// TIA Portal project "FORMING_1500_PLC" (V15) (continued)
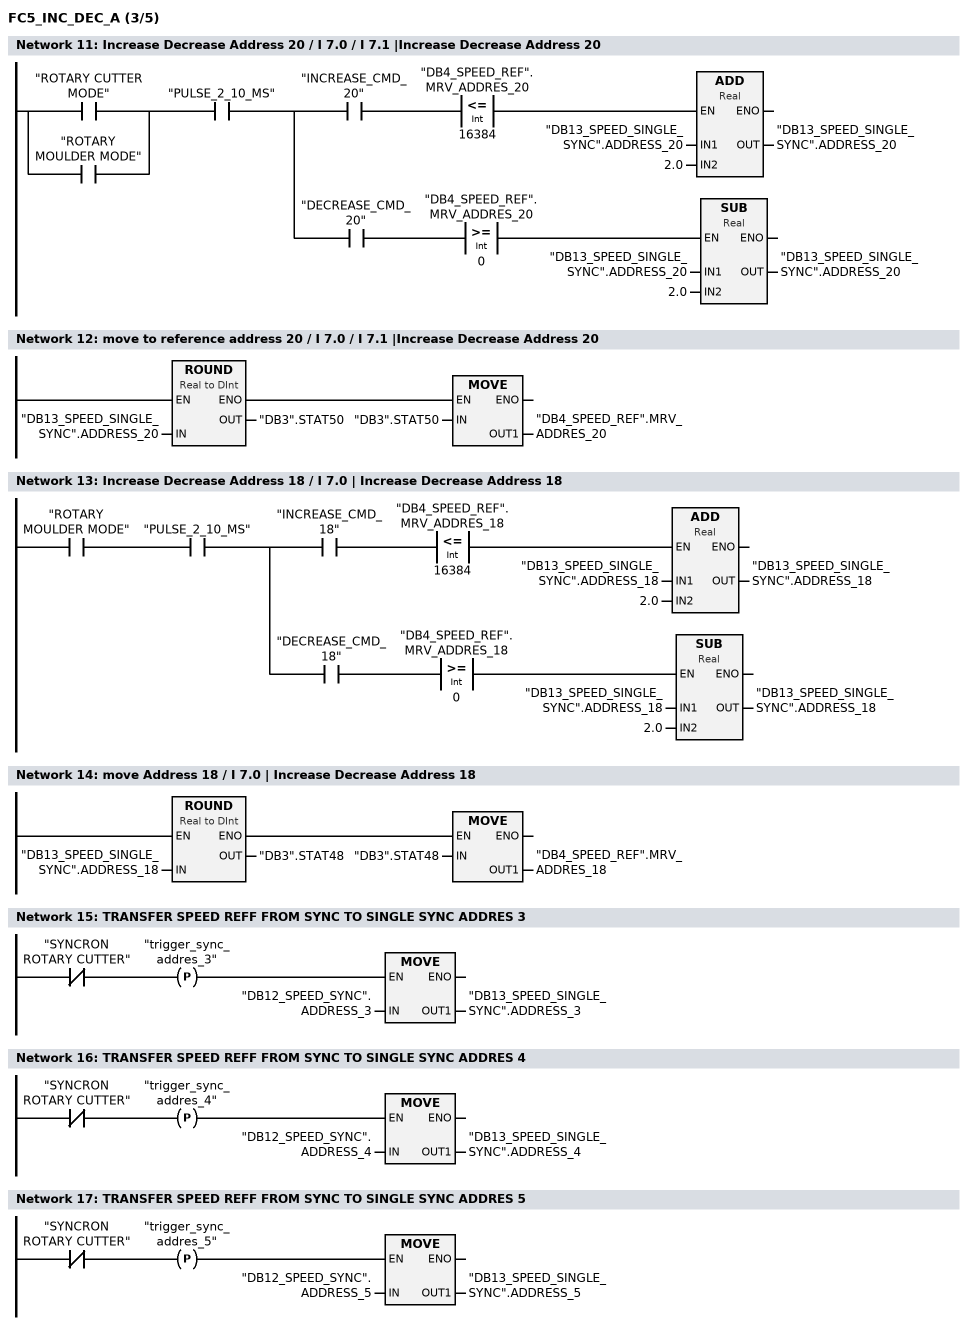
   RUNG wire#powerrail
      Contact( "ROTARY CUTTER MODE" )
      wire#w1
      Contact( "PULSE_2_10_MS" )
      wire#w2
      Contact( "INCREASE_CMD_20" )
      { S7_Templates := "SrcType := Int" } LE_Contact(in1 := "DB4_SPEED_REF".MRV_ADDRES_20, in2 := 16384)
      { S7_Templates := "SrcType := Real"; S7_GenerateENO := "TRUE" } Add(in1 := "DB13_SPEED_SINGLE_SYNC".ADDRESS_20, in2 := 2.0, out => "DB13_SPEED_SINGLE_SYNC".ADDRESS_20)
   END_RUNG
   RUNG wire#powerrail
      Contact( "ROTARY MOULDER MODE" )
   END_RUNG wire#w1
   RUNG wire#w2
      Contact( "DECREASE_CMD_20" )
      { S7_Templates := "SrcType := Int" } GE_Contact(in1 := "DB4_SPEED_REF".MRV_ADDRES_20, in2 := 0)
      { S7_Templates := "SrcType := Real"; S7_GenerateENO := "TRUE" } Sub(in1 := "DB13_SPEED_SINGLE_SYNC".ADDRESS_20, in2 := 2.0, out => "DB13_SPEED_SINGLE_SYNC".ADDRESS_20)
   END_RUNG
   // the same network as SCL:
   #_w1 := ("ROTARY CUTTER MODE" OR "ROTARY MOULDER MODE") AND "PULSE_2_10_MS";
   IF #_w1 AND "INCREASE_CMD_20" AND ("DB4_SPEED_REF".MRV_ADDRES_20 <= 16384) THEN
       "DB13_SPEED_SINGLE_SYNC".ADDRESS_20 := "DB13_SPEED_SINGLE_SYNC".ADDRESS_20 + 2.0;
   END_IF;
   IF #_w1 AND "DECREASE_CMD_20" AND ("DB4_SPEED_REF".MRV_ADDRES_20 >= 0) THEN
       "DB13_SPEED_SINGLE_SYNC".ADDRESS_20 := "DB13_SPEED_SINGLE_SYNC".ADDRESS_20 - 2.0;
   END_IF;
END_REGION

REGION Network 12: move to reference address 20 / I 7.0 / I 7.1 |Increase Decrease Address 20
   RUNG wire#powerrail
      { S7_Templates := "[SrcType := Real, DestType := DInt]"; S7_GenerateENO := "TRUE" } Round(in := "DB13_SPEED_SINGLE_SYNC".ADDRESS_20, out => "DB3".STAT50)
      { S7_GenerateENO := "TRUE" } Move(in := "DB3".STAT50, out1 => "DB4_SPEED_REF".MRV_ADDRES_20)
   END_RUNG
   // the same network as SCL:
   // ENO of a box is taken as its EN; it also drops when the box reports an error
   "DB3".STAT50 := ROUND("DB13_SPEED_SINGLE_SYNC".ADDRESS_20);
   "DB4_SPEED_REF".MRV_ADDRES_20 := "DB3".STAT50;
END_REGION

REGION Network 13: Increase Decrease Address 18 / I 7.0 | Increase Decrease Address 18
   RUNG wire#powerrail
      Contact( "ROTARY MOULDER MODE" )
      Contact( "PULSE_2_10_MS" )
      wire#w1
      Contact( "INCREASE_CMD_18" )
      { S7_Templates := "SrcType := Int" } LE_Contact(in1 := "DB4_SPEED_REF".MRV_ADDRES_18, in2 := 16384)
      { S7_Templates := "SrcType := Real"; S7_GenerateENO := "TRUE" } Add(in1 := "DB13_SPEED_SINGLE_SYNC".ADDRESS_18, in2 := 2.0, out => "DB13_SPEED_SINGLE_SYNC".ADDRESS_18)
   END_RUNG
   RUNG wire#w1
      Contact( "DECREASE_CMD_18" )
      { S7_Templates := "SrcType := Int" } GE_Contact(in1 := "DB4_SPEED_REF".MRV_ADDRES_18, in2 := 0)
      { S7_Templates := "SrcType := Real"; S7_GenerateENO := "TRUE" } Sub(in1 := "DB13_SPEED_SINGLE_SYNC".ADDRESS_18, in2 := 2.0, out => "DB13_SPEED_SINGLE_SYNC".ADDRESS_18)
   END_RUNG
   // the same network as SCL:
   #_w1 := "ROTARY MOULDER MODE" AND "PULSE_2_10_MS";
   IF #_w1 AND "INCREASE_CMD_18" AND ("DB4_SPEED_REF".MRV_ADDRES_18 <= 16384) THEN
       "DB13_SPEED_SINGLE_SYNC".ADDRESS_18 := "DB13_SPEED_SINGLE_SYNC".ADDRESS_18 + 2.0;
   END_IF;
   IF #_w1 AND "DECREASE_CMD_18" AND ("DB4_SPEED_REF".MRV_ADDRES_18 >= 0) THEN
       "DB13_SPEED_SINGLE_SYNC".ADDRESS_18 := "DB13_SPEED_SINGLE_SYNC".ADDRESS_18 - 2.0;
   END_IF;
END_REGION

REGION Network 14: move Address 18 / I 7.0 | Increase Decrease Address 18
   RUNG wire#powerrail
      { S7_Templates := "[SrcType := Real, DestType := DInt]"; S7_GenerateENO := "TRUE" } Round(in := "DB13_SPEED_SINGLE_SYNC".ADDRESS_18, out => "DB3".STAT48)
      { S7_GenerateENO := "TRUE" } Move(in := "DB3".STAT48, out1 => "DB4_SPEED_REF".MRV_ADDRES_18)
   END_RUNG
   // the same network as SCL:
   // ENO of a box is taken as its EN; it also drops when the box reports an error
   "DB3".STAT48 := ROUND("DB13_SPEED_SINGLE_SYNC".ADDRESS_18);
   "DB4_SPEED_REF".MRV_ADDRES_18 := "DB3".STAT48;
END_REGION

REGION Network 15: TRANSFER SPEED REFF FROM SYNC TO SINGLE SYNC ADDRES 3
   RUNG wire#powerrail
      I_Contact( "SYNCRON ROTARY CUTTER" )
      P_Trig( "trigger_sync_addres_3" )
      { S7_GenerateENO := "TRUE" } Move(in := "DB12_SPEED_SYNC".ADDRESS_3, out1 => "DB13_SPEED_SINGLE_SYNC".ADDRESS_3)
   END_RUNG
   // the same network as SCL:
   #_w1 := NOT "SYNCRON ROTARY CUTTER" AND NOT "trigger_sync_addres_3";   // rising edge
   "trigger_sync_addres_3" := NOT "SYNCRON ROTARY CUTTER";
   IF #_w1 THEN "DB13_SPEED_SINGLE_SYNC".ADDRESS_3 := "DB12_SPEED_SYNC".ADDRESS_3; END_IF;
END_REGION

REGION Network 16: TRANSFER SPEED REFF FROM SYNC TO SINGLE SYNC ADDRES 4
   RUNG wire#powerrail
      I_Contact( "SYNCRON ROTARY CUTTER" )
      P_Trig( "trigger_sync_addres_4" )
      { S7_GenerateENO := "TRUE" } Move(in := "DB12_SPEED_SYNC".ADDRESS_4, out1 => "DB13_SPEED_SINGLE_SYNC".ADDRESS_4)
   END_RUNG
   // the same network as SCL:
   #_w1 := NOT "SYNCRON ROTARY CUTTER" AND NOT "trigger_sync_addres_4";   // rising edge
   "trigger_sync_addres_4" := NOT "SYNCRON ROTARY CUTTER";
   IF #_w1 THEN "DB13_SPEED_SINGLE_SYNC".ADDRESS_4 := "DB12_SPEED_SYNC".ADDRESS_4; END_IF;
END_REGION

REGION Network 17: TRANSFER SPEED REFF FROM SYNC TO SINGLE SYNC ADDRES 5
   RUNG wire#powerrail
      I_Contact( "SYNCRON ROTARY CUTTER" )
      P_Trig( "trigger_sync_addres_5" )
      { S7_GenerateENO := "TRUE" } Move(in := "DB12_SPEED_SYNC".ADDRESS_5, out1 => "DB13_SPEED_SINGLE_SYNC".ADDRESS_5)
   END_RUNG
   // the same network as SCL:
   #_w1 := NOT "SYNCRON ROTARY CUTTER" AND NOT "trigger_sync_addres_5";   // rising edge
   "trigger_sync_addres_5" := NOT "SYNCRON ROTARY CUTTER";
   IF #_w1 THEN "DB13_SPEED_SINGLE_SYNC".ADDRESS_5 := "DB12_SPEED_SYNC".ADDRESS_5; END_IF;
END_REGION

REGION Network 18: TRANSFER SPEED REFF FROM SYNC TO SINGLE SYNC ADDRES 6
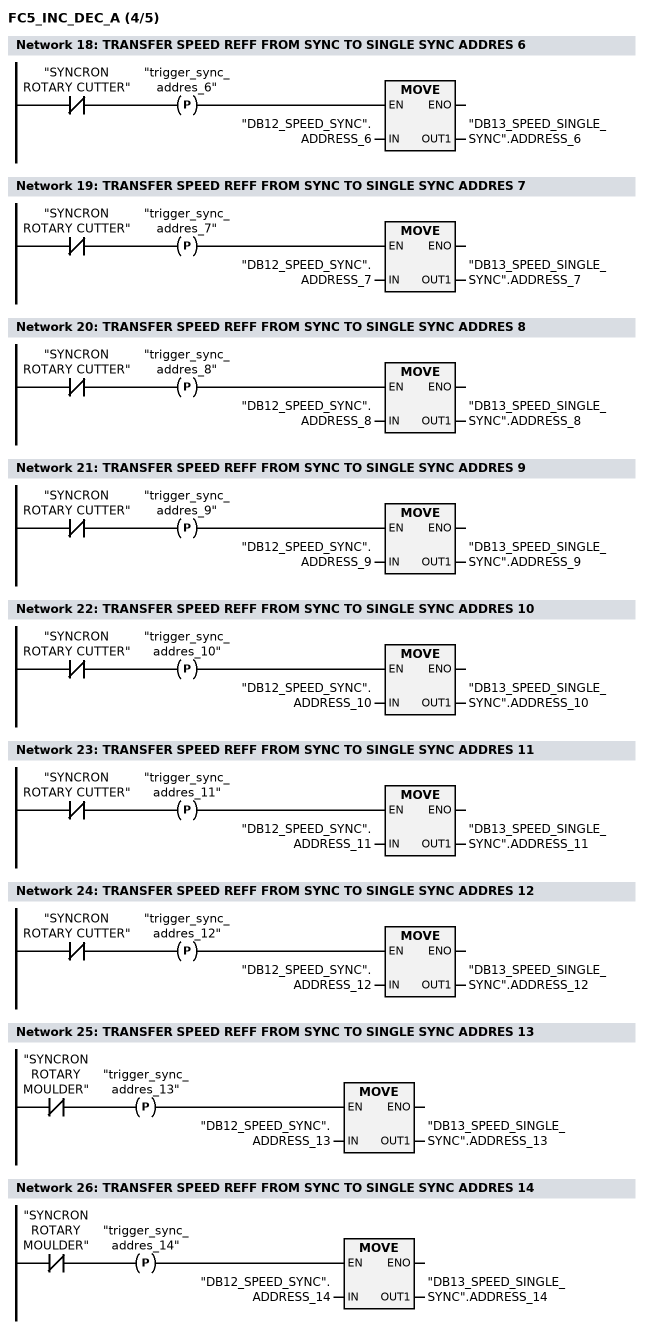
   RUNG wire#powerrail
      I_Contact( "SYNCRON ROTARY CUTTER" )
      P_Trig( "trigger_sync_addres_6" )
      { S7_GenerateENO := "TRUE" } Move(in := "DB12_SPEED_SYNC".ADDRESS_6, out1 => "DB13_SPEED_SINGLE_SYNC".ADDRESS_6)
   END_RUNG
   // the same network as SCL:
   #_w1 := NOT "SYNCRON ROTARY CUTTER" AND NOT "trigger_sync_addres_6";   // rising edge
   "trigger_sync_addres_6" := NOT "SYNCRON ROTARY CUTTER";
   IF #_w1 THEN "DB13_SPEED_SINGLE_SYNC".ADDRESS_6 := "DB12_SPEED_SYNC".ADDRESS_6; END_IF;
END_REGION

REGION Network 19: TRANSFER SPEED REFF FROM SYNC TO SINGLE SYNC ADDRES 7
   RUNG wire#powerrail
      I_Contact( "SYNCRON ROTARY CUTTER" )
      P_Trig( "trigger_sync_addres_7" )
      { S7_GenerateENO := "TRUE" } Move(in := "DB12_SPEED_SYNC".ADDRESS_7, out1 => "DB13_SPEED_SINGLE_SYNC".ADDRESS_7)
   END_RUNG
   // the same network as SCL:
   #_w1 := NOT "SYNCRON ROTARY CUTTER" AND NOT "trigger_sync_addres_7";   // rising edge
   "trigger_sync_addres_7" := NOT "SYNCRON ROTARY CUTTER";
   IF #_w1 THEN "DB13_SPEED_SINGLE_SYNC".ADDRESS_7 := "DB12_SPEED_SYNC".ADDRESS_7; END_IF;
END_REGION

REGION Network 20: TRANSFER SPEED REFF FROM SYNC TO SINGLE SYNC ADDRES 8
   RUNG wire#powerrail
      I_Contact( "SYNCRON ROTARY CUTTER" )
      P_Trig( "trigger_sync_addres_8" )
      { S7_GenerateENO := "TRUE" } Move(in := "DB12_SPEED_SYNC".ADDRESS_8, out1 => "DB13_SPEED_SINGLE_SYNC".ADDRESS_8)
   END_RUNG
   // the same network as SCL:
   #_w1 := NOT "SYNCRON ROTARY CUTTER" AND NOT "trigger_sync_addres_8";   // rising edge
   "trigger_sync_addres_8" := NOT "SYNCRON ROTARY CUTTER";
   IF #_w1 THEN "DB13_SPEED_SINGLE_SYNC".ADDRESS_8 := "DB12_SPEED_SYNC".ADDRESS_8; END_IF;
END_REGION

REGION Network 21: TRANSFER SPEED REFF FROM SYNC TO SINGLE SYNC ADDRES 9
   RUNG wire#powerrail
      I_Contact( "SYNCRON ROTARY CUTTER" )
      P_Trig( "trigger_sync_addres_9" )
      { S7_GenerateENO := "TRUE" } Move(in := "DB12_SPEED_SYNC".ADDRESS_9, out1 => "DB13_SPEED_SINGLE_SYNC".ADDRESS_9)
   END_RUNG
   // the same network as SCL:
   #_w1 := NOT "SYNCRON ROTARY CUTTER" AND NOT "trigger_sync_addres_9";   // rising edge
   "trigger_sync_addres_9" := NOT "SYNCRON ROTARY CUTTER";
   IF #_w1 THEN "DB13_SPEED_SINGLE_SYNC".ADDRESS_9 := "DB12_SPEED_SYNC".ADDRESS_9; END_IF;
END_REGION

REGION Network 22: TRANSFER SPEED REFF FROM SYNC TO SINGLE SYNC ADDRES 10
   RUNG wire#powerrail
      I_Contact( "SYNCRON ROTARY CUTTER" )
      P_Trig( "trigger_sync_addres_10" )
      { S7_GenerateENO := "TRUE" } Move(in := "DB12_SPEED_SYNC".ADDRESS_10, out1 => "DB13_SPEED_SINGLE_SYNC".ADDRESS_10)
   END_RUNG
   // the same network as SCL:
   #_w1 := NOT "SYNCRON ROTARY CUTTER" AND NOT "trigger_sync_addres_10";   // rising edge
   "trigger_sync_addres_10" := NOT "SYNCRON ROTARY CUTTER";
   IF #_w1 THEN "DB13_SPEED_SINGLE_SYNC".ADDRESS_10 := "DB12_SPEED_SYNC".ADDRESS_10; END_IF;
END_REGION

REGION Network 23: TRANSFER SPEED REFF FROM SYNC TO SINGLE SYNC ADDRES 11
   RUNG wire#powerrail
      I_Contact( "SYNCRON ROTARY CUTTER" )
      P_Trig( "trigger_sync_addres_11" )
      { S7_GenerateENO := "TRUE" } Move(in := "DB12_SPEED_SYNC".ADDRESS_11, out1 => "DB13_SPEED_SINGLE_SYNC".ADDRESS_11)
   END_RUNG
   // the same network as SCL:
   #_w1 := NOT "SYNCRON ROTARY CUTTER" AND NOT "trigger_sync_addres_11";   // rising edge
   "trigger_sync_addres_11" := NOT "SYNCRON ROTARY CUTTER";
   IF #_w1 THEN "DB13_SPEED_SINGLE_SYNC".ADDRESS_11 := "DB12_SPEED_SYNC".ADDRESS_11; END_IF;
END_REGION

REGION Network 24: TRANSFER SPEED REFF FROM SYNC TO SINGLE SYNC ADDRES 12
   RUNG wire#powerrail
      I_Contact( "SYNCRON ROTARY CUTTER" )
      P_Trig( "trigger_sync_addres_12" )
      { S7_GenerateENO := "TRUE" } Move(in := "DB12_SPEED_SYNC".ADDRESS_12, out1 => "DB13_SPEED_SINGLE_SYNC".ADDRESS_12)
   END_RUNG
   // the same network as SCL:
   #_w1 := NOT "SYNCRON ROTARY CUTTER" AND NOT "trigger_sync_addres_12";   // rising edge
   "trigger_sync_addres_12" := NOT "SYNCRON ROTARY CUTTER";
   IF #_w1 THEN "DB13_SPEED_SINGLE_SYNC".ADDRESS_12 := "DB12_SPEED_SYNC".ADDRESS_12; END_IF;
END_REGION

REGION Network 25: TRANSFER SPEED REFF FROM SYNC TO SINGLE SYNC ADDRES 13
   RUNG wire#powerrail
      I_Contact( "SYNCRON ROTARY MOULDER" )
      P_Trig( "trigger_sync_addres_13" )
      { S7_GenerateENO := "TRUE" } Move(in := "DB12_SPEED_SYNC".ADDRESS_13, out1 => "DB13_SPEED_SINGLE_SYNC".ADDRESS_13)
   END_RUNG
   // the same network as SCL:
   #_w1 := NOT "SYNCRON ROTARY MOULDER" AND NOT "trigger_sync_addres_13";   // rising edge
   "trigger_sync_addres_13" := NOT "SYNCRON ROTARY MOULDER";
   IF #_w1 THEN "DB13_SPEED_SINGLE_SYNC".ADDRESS_13 := "DB12_SPEED_SYNC".ADDRESS_13; END_IF;
END_REGION

REGION Network 26: TRANSFER SPEED REFF FROM SYNC TO SINGLE SYNC ADDRES 14
   RUNG wire#powerrail
      I_Contact( "SYNCRON ROTARY MOULDER" )
      P_Trig( "trigger_sync_addres_14" )
      { S7_GenerateENO := "TRUE" } Move(in := "DB12_SPEED_SYNC".ADDRESS_14, out1 => "DB13_SPEED_SINGLE_SYNC".ADDRESS_14)
   END_RUNG
   // the same network as SCL:
   #_w1 := NOT "SYNCRON ROTARY MOULDER" AND NOT "trigger_sync_addres_14";   // rising edge
   "trigger_sync_addres_14" := NOT "SYNCRON ROTARY MOULDER";
   IF #_w1 THEN "DB13_SPEED_SINGLE_SYNC".ADDRESS_14 := "DB12_SPEED_SYNC".ADDRESS_14; END_IF;
END_REGION

REGION Network 27: TRANSFER SPEED REFF FROM SYNC TO SINGLE SYNC ADDRES 15
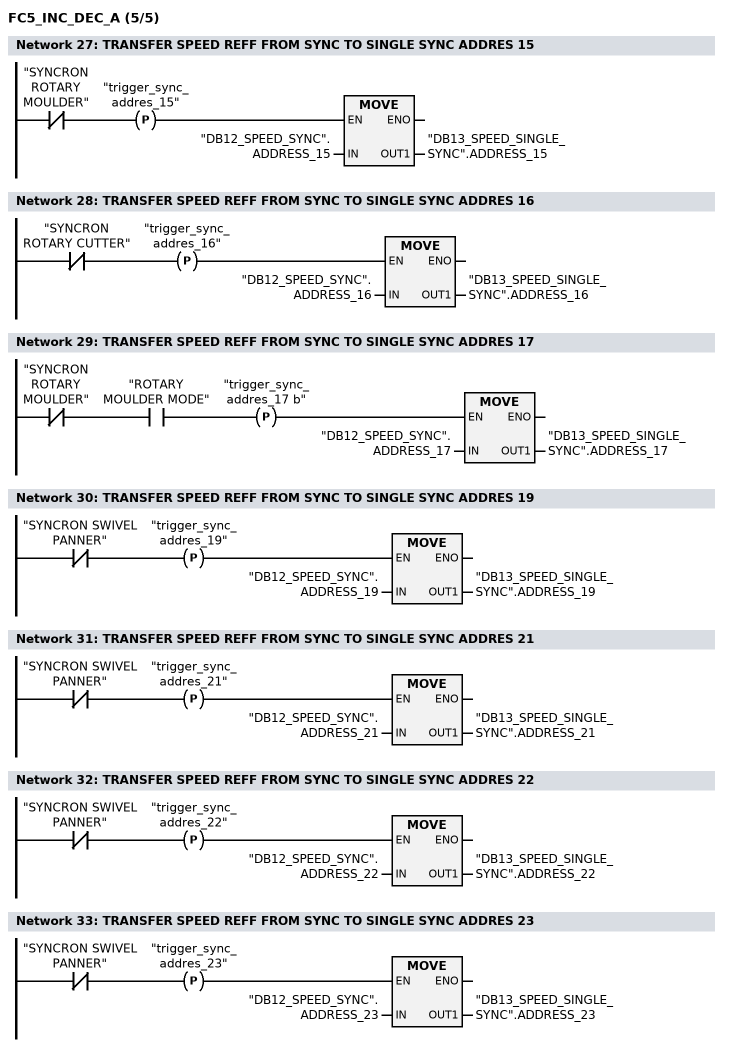
   RUNG wire#powerrail
      I_Contact( "SYNCRON ROTARY MOULDER" )
      P_Trig( "trigger_sync_addres_15" )
      { S7_GenerateENO := "TRUE" } Move(in := "DB12_SPEED_SYNC".ADDRESS_15, out1 => "DB13_SPEED_SINGLE_SYNC".ADDRESS_15)
   END_RUNG
   // the same network as SCL:
   #_w1 := NOT "SYNCRON ROTARY MOULDER" AND NOT "trigger_sync_addres_15";   // rising edge
   "trigger_sync_addres_15" := NOT "SYNCRON ROTARY MOULDER";
   IF #_w1 THEN "DB13_SPEED_SINGLE_SYNC".ADDRESS_15 := "DB12_SPEED_SYNC".ADDRESS_15; END_IF;
END_REGION

REGION Network 28: TRANSFER SPEED REFF FROM SYNC TO SINGLE SYNC ADDRES 16
   RUNG wire#powerrail
      I_Contact( "SYNCRON ROTARY CUTTER" )
      P_Trig( "trigger_sync_addres_16" )
      { S7_GenerateENO := "TRUE" } Move(in := "DB12_SPEED_SYNC".ADDRESS_16, out1 => "DB13_SPEED_SINGLE_SYNC".ADDRESS_16)
   END_RUNG
   // the same network as SCL:
   #_w1 := NOT "SYNCRON ROTARY CUTTER" AND NOT "trigger_sync_addres_16";   // rising edge
   "trigger_sync_addres_16" := NOT "SYNCRON ROTARY CUTTER";
   IF #_w1 THEN "DB13_SPEED_SINGLE_SYNC".ADDRESS_16 := "DB12_SPEED_SYNC".ADDRESS_16; END_IF;
END_REGION

REGION Network 29: TRANSFER SPEED REFF FROM SYNC TO SINGLE SYNC ADDRES 17
   RUNG wire#powerrail
      I_Contact( "SYNCRON ROTARY MOULDER" )
      Contact( "ROTARY MOULDER MODE" )
      P_Trig( "trigger_sync_addres_17 b" )
      { S7_GenerateENO := "TRUE" } Move(in := "DB12_SPEED_SYNC".ADDRESS_17, out1 => "DB13_SPEED_SINGLE_SYNC".ADDRESS_17)
   END_RUNG
   // the same network as SCL:
   #_w1 := NOT "SYNCRON ROTARY MOULDER" AND "ROTARY MOULDER MODE";
   #_w2 := #_w1 AND NOT "trigger_sync_addres_17 b";   // rising edge
   "trigger_sync_addres_17 b" := #_w1;
   IF #_w2 THEN "DB13_SPEED_SINGLE_SYNC".ADDRESS_17 := "DB12_SPEED_SYNC".ADDRESS_17; END_IF;
END_REGION

REGION Network 30: TRANSFER SPEED REFF FROM SYNC TO SINGLE SYNC ADDRES 19
   RUNG wire#powerrail
      I_Contact( "SYNCRON SWIVEL PANNER" )
      P_Trig( "trigger_sync_addres_19" )
      { S7_GenerateENO := "TRUE" } Move(in := "DB12_SPEED_SYNC".ADDRESS_19, out1 => "DB13_SPEED_SINGLE_SYNC".ADDRESS_19)
   END_RUNG
   // the same network as SCL:
   #_w1 := NOT "SYNCRON SWIVEL PANNER" AND NOT "trigger_sync_addres_19";   // rising edge
   "trigger_sync_addres_19" := NOT "SYNCRON SWIVEL PANNER";
   IF #_w1 THEN "DB13_SPEED_SINGLE_SYNC".ADDRESS_19 := "DB12_SPEED_SYNC".ADDRESS_19; END_IF;
END_REGION

REGION Network 31: TRANSFER SPEED REFF FROM SYNC TO SINGLE SYNC ADDRES 21
   RUNG wire#powerrail
      I_Contact( "SYNCRON SWIVEL PANNER" )
      P_Trig( "trigger_sync_addres_21" )
      { S7_GenerateENO := "TRUE" } Move(in := "DB12_SPEED_SYNC".ADDRESS_21, out1 => "DB13_SPEED_SINGLE_SYNC".ADDRESS_21)
   END_RUNG
   // the same network as SCL:
   #_w1 := NOT "SYNCRON SWIVEL PANNER" AND NOT "trigger_sync_addres_21";   // rising edge
   "trigger_sync_addres_21" := NOT "SYNCRON SWIVEL PANNER";
   IF #_w1 THEN "DB13_SPEED_SINGLE_SYNC".ADDRESS_21 := "DB12_SPEED_SYNC".ADDRESS_21; END_IF;
END_REGION

REGION Network 32: TRANSFER SPEED REFF FROM SYNC TO SINGLE SYNC ADDRES 22
   RUNG wire#powerrail
      I_Contact( "SYNCRON SWIVEL PANNER" )
      P_Trig( "trigger_sync_addres_22" )
      { S7_GenerateENO := "TRUE" } Move(in := "DB12_SPEED_SYNC".ADDRESS_22, out1 => "DB13_SPEED_SINGLE_SYNC".ADDRESS_22)
   END_RUNG
   // the same network as SCL:
   #_w1 := NOT "SYNCRON SWIVEL PANNER" AND NOT "trigger_sync_addres_22";   // rising edge
   "trigger_sync_addres_22" := NOT "SYNCRON SWIVEL PANNER";
   IF #_w1 THEN "DB13_SPEED_SINGLE_SYNC".ADDRESS_22 := "DB12_SPEED_SYNC".ADDRESS_22; END_IF;
END_REGION

REGION Network 33: TRANSFER SPEED REFF FROM SYNC TO SINGLE SYNC ADDRES 23
   RUNG wire#powerrail
      I_Contact( "SYNCRON SWIVEL PANNER" )
      P_Trig( "trigger_sync_addres_23" )
      { S7_GenerateENO := "TRUE" } Move(in := "DB12_SPEED_SYNC".ADDRESS_23, out1 => "DB13_SPEED_SINGLE_SYNC".ADDRESS_23)
   END_RUNG
   // the same network as SCL:
   #_w1 := NOT "SYNCRON SWIVEL PANNER" AND NOT "trigger_sync_addres_23";   // rising edge
   "trigger_sync_addres_23" := NOT "SYNCRON SWIVEL PANNER";
   IF #_w1 THEN "DB13_SPEED_SINGLE_SYNC".ADDRESS_23 := "DB12_SPEED_SYNC".ADDRESS_23; END_IF;
END_REGION
END_FUNCTION

FUNCTION "FC6_SPEED ACTUAL / MAV" : Void   // FC6, LAD
TITLE = MAIN ACTUAL VALUE DARI INVERTER VLT
{ S7_Optimized_Access := 'FALSE' }
VERSION : 0.1
BEGIN

REGION Network 1: MAIN ACTUAL VALUE / FEEDBACK SPEED ADDRES 2
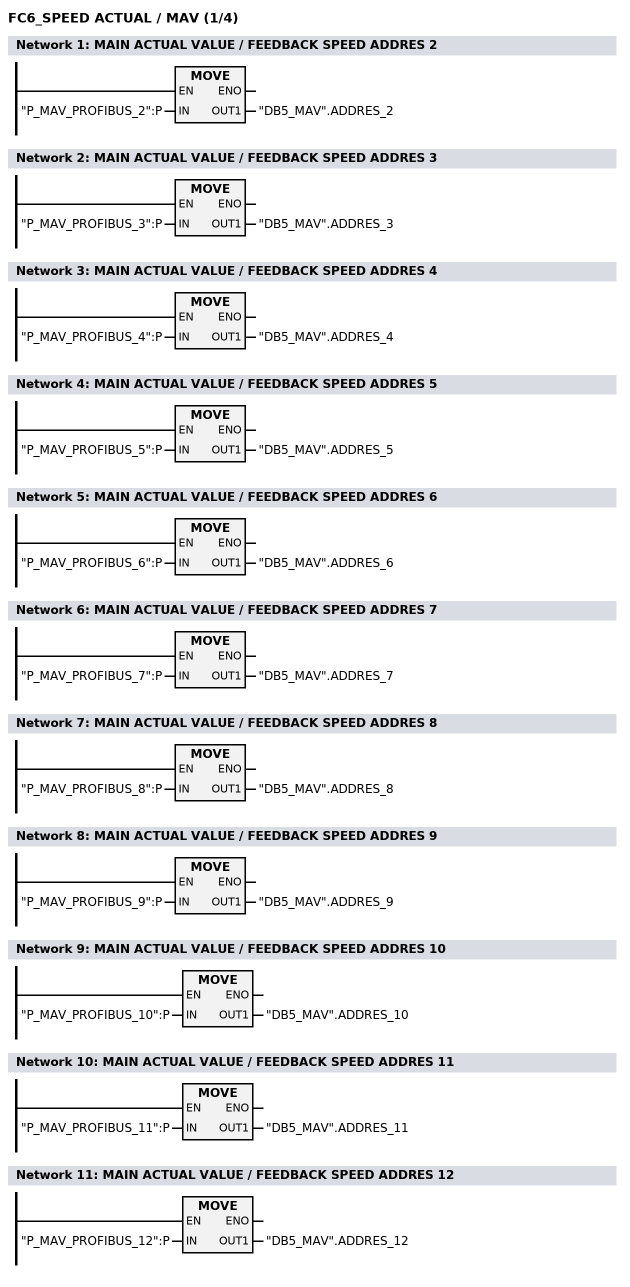
   RUNG wire#powerrail
      { S7_GenerateENO := "TRUE" } Move(in := "P_MAV_PROFIBUS_2":P, out1 => "DB5_MAV".ADDRES_2)
   END_RUNG
   // the same network as SCL:
   "DB5_MAV".ADDRES_2 := "P_MAV_PROFIBUS_2":P;
END_REGION

REGION Network 2: MAIN ACTUAL VALUE / FEEDBACK SPEED ADDRES 3
   RUNG wire#powerrail
      { S7_GenerateENO := "TRUE" } Move(in := "P_MAV_PROFIBUS_3":P, out1 => "DB5_MAV".ADDRES_3)
   END_RUNG
   // the same network as SCL:
   "DB5_MAV".ADDRES_3 := "P_MAV_PROFIBUS_3":P;
END_REGION

REGION Network 3: MAIN ACTUAL VALUE / FEEDBACK SPEED ADDRES 4
   RUNG wire#powerrail
      { S7_GenerateENO := "TRUE" } Move(in := "P_MAV_PROFIBUS_4":P, out1 => "DB5_MAV".ADDRES_4)
   END_RUNG
   // the same network as SCL:
   "DB5_MAV".ADDRES_4 := "P_MAV_PROFIBUS_4":P;
END_REGION

REGION Network 4: MAIN ACTUAL VALUE / FEEDBACK SPEED ADDRES 5
   RUNG wire#powerrail
      { S7_GenerateENO := "TRUE" } Move(in := "P_MAV_PROFIBUS_5":P, out1 => "DB5_MAV".ADDRES_5)
   END_RUNG
   // the same network as SCL:
   "DB5_MAV".ADDRES_5 := "P_MAV_PROFIBUS_5":P;
END_REGION

REGION Network 5: MAIN ACTUAL VALUE / FEEDBACK SPEED ADDRES 6
   RUNG wire#powerrail
      { S7_GenerateENO := "TRUE" } Move(in := "P_MAV_PROFIBUS_6":P, out1 => "DB5_MAV".ADDRES_6)
   END_RUNG
   // the same network as SCL:
   "DB5_MAV".ADDRES_6 := "P_MAV_PROFIBUS_6":P;
END_REGION

REGION Network 6: MAIN ACTUAL VALUE / FEEDBACK SPEED ADDRES 7
   RUNG wire#powerrail
      { S7_GenerateENO := "TRUE" } Move(in := "P_MAV_PROFIBUS_7":P, out1 => "DB5_MAV".ADDRES_7)
   END_RUNG
   // the same network as SCL:
   "DB5_MAV".ADDRES_7 := "P_MAV_PROFIBUS_7":P;
END_REGION

REGION Network 7: MAIN ACTUAL VALUE / FEEDBACK SPEED ADDRES 8
   RUNG wire#powerrail
      { S7_GenerateENO := "TRUE" } Move(in := "P_MAV_PROFIBUS_8":P, out1 => "DB5_MAV".ADDRES_8)
   END_RUNG
   // the same network as SCL:
   "DB5_MAV".ADDRES_8 := "P_MAV_PROFIBUS_8":P;
END_REGION

REGION Network 8: MAIN ACTUAL VALUE / FEEDBACK SPEED ADDRES 9
   RUNG wire#powerrail
      { S7_GenerateENO := "TRUE" } Move(in := "P_MAV_PROFIBUS_9":P, out1 => "DB5_MAV".ADDRES_9)
   END_RUNG
   // the same network as SCL:
   "DB5_MAV".ADDRES_9 := "P_MAV_PROFIBUS_9":P;
END_REGION

REGION Network 9: MAIN ACTUAL VALUE / FEEDBACK SPEED ADDRES 10
   RUNG wire#powerrail
      { S7_GenerateENO := "TRUE" } Move(in := "P_MAV_PROFIBUS_10":P, out1 => "DB5_MAV".ADDRES_10)
   END_RUNG
   // the same network as SCL:
   "DB5_MAV".ADDRES_10 := "P_MAV_PROFIBUS_10":P;
END_REGION

REGION Network 10: MAIN ACTUAL VALUE / FEEDBACK SPEED ADDRES 11
   RUNG wire#powerrail
      { S7_GenerateENO := "TRUE" } Move(in := "P_MAV_PROFIBUS_11":P, out1 => "DB5_MAV".ADDRES_11)
   END_RUNG
   // the same network as SCL:
   "DB5_MAV".ADDRES_11 := "P_MAV_PROFIBUS_11":P;
END_REGION

REGION Network 11: MAIN ACTUAL VALUE / FEEDBACK SPEED ADDRES 12
   RUNG wire#powerrail
      { S7_GenerateENO := "TRUE" } Move(in := "P_MAV_PROFIBUS_12":P, out1 => "DB5_MAV".ADDRES_12)
   END_RUNG
   // the same network as SCL:
   "DB5_MAV".ADDRES_12 := "P_MAV_PROFIBUS_12":P;
END_REGION

REGION Network 12: MAIN ACTUAL VALUE / FEEDBACK SPEED ADDRES 13
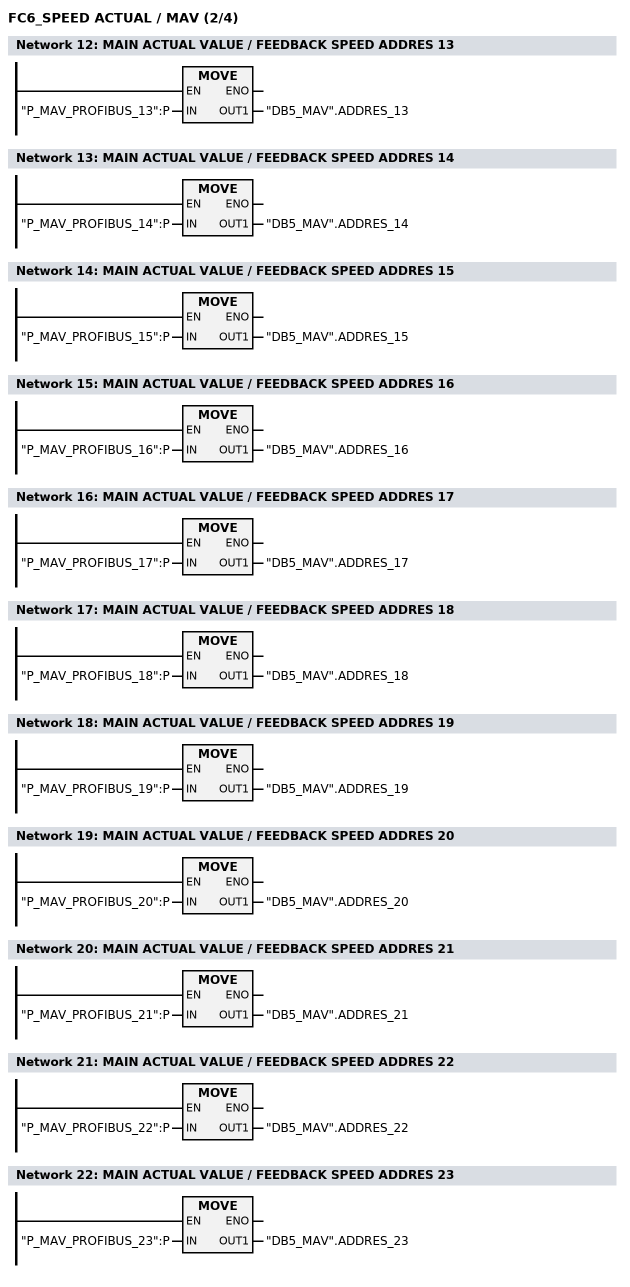
   RUNG wire#powerrail
      { S7_GenerateENO := "TRUE" } Move(in := "P_MAV_PROFIBUS_13":P, out1 => "DB5_MAV".ADDRES_13)
   END_RUNG
   // the same network as SCL:
   "DB5_MAV".ADDRES_13 := "P_MAV_PROFIBUS_13":P;
END_REGION

REGION Network 13: MAIN ACTUAL VALUE / FEEDBACK SPEED ADDRES 14
   RUNG wire#powerrail
      { S7_GenerateENO := "TRUE" } Move(in := "P_MAV_PROFIBUS_14":P, out1 => "DB5_MAV".ADDRES_14)
   END_RUNG
   // the same network as SCL:
   "DB5_MAV".ADDRES_14 := "P_MAV_PROFIBUS_14":P;
END_REGION

REGION Network 14: MAIN ACTUAL VALUE / FEEDBACK SPEED ADDRES 15
   RUNG wire#powerrail
      { S7_GenerateENO := "TRUE" } Move(in := "P_MAV_PROFIBUS_15":P, out1 => "DB5_MAV".ADDRES_15)
   END_RUNG
   // the same network as SCL:
   "DB5_MAV".ADDRES_15 := "P_MAV_PROFIBUS_15":P;
END_REGION

REGION Network 15: MAIN ACTUAL VALUE / FEEDBACK SPEED ADDRES 16
   RUNG wire#powerrail
      { S7_GenerateENO := "TRUE" } Move(in := "P_MAV_PROFIBUS_16":P, out1 => "DB5_MAV".ADDRES_16)
   END_RUNG
   // the same network as SCL:
   "DB5_MAV".ADDRES_16 := "P_MAV_PROFIBUS_16":P;
END_REGION

REGION Network 16: MAIN ACTUAL VALUE / FEEDBACK SPEED ADDRES 17
   RUNG wire#powerrail
      { S7_GenerateENO := "TRUE" } Move(in := "P_MAV_PROFIBUS_17":P, out1 => "DB5_MAV".ADDRES_17)
   END_RUNG
   // the same network as SCL:
   "DB5_MAV".ADDRES_17 := "P_MAV_PROFIBUS_17":P;
END_REGION

REGION Network 17: MAIN ACTUAL VALUE / FEEDBACK SPEED ADDRES 18
   RUNG wire#powerrail
      { S7_GenerateENO := "TRUE" } Move(in := "P_MAV_PROFIBUS_18":P, out1 => "DB5_MAV".ADDRES_18)
   END_RUNG
   // the same network as SCL:
   "DB5_MAV".ADDRES_18 := "P_MAV_PROFIBUS_18":P;
END_REGION

REGION Network 18: MAIN ACTUAL VALUE / FEEDBACK SPEED ADDRES 19
   RUNG wire#powerrail
      { S7_GenerateENO := "TRUE" } Move(in := "P_MAV_PROFIBUS_19":P, out1 => "DB5_MAV".ADDRES_19)
   END_RUNG
   // the same network as SCL:
   "DB5_MAV".ADDRES_19 := "P_MAV_PROFIBUS_19":P;
END_REGION

REGION Network 19: MAIN ACTUAL VALUE / FEEDBACK SPEED ADDRES 20
   RUNG wire#powerrail
      { S7_GenerateENO := "TRUE" } Move(in := "P_MAV_PROFIBUS_20":P, out1 => "DB5_MAV".ADDRES_20)
   END_RUNG
   // the same network as SCL:
   "DB5_MAV".ADDRES_20 := "P_MAV_PROFIBUS_20":P;
END_REGION

REGION Network 20: MAIN ACTUAL VALUE / FEEDBACK SPEED ADDRES 21
   RUNG wire#powerrail
      { S7_GenerateENO := "TRUE" } Move(in := "P_MAV_PROFIBUS_21":P, out1 => "DB5_MAV".ADDRES_21)
   END_RUNG
   // the same network as SCL:
   "DB5_MAV".ADDRES_21 := "P_MAV_PROFIBUS_21":P;
END_REGION

REGION Network 21: MAIN ACTUAL VALUE / FEEDBACK SPEED ADDRES 22
   RUNG wire#powerrail
      { S7_GenerateENO := "TRUE" } Move(in := "P_MAV_PROFIBUS_22":P, out1 => "DB5_MAV".ADDRES_22)
   END_RUNG
   // the same network as SCL:
   "DB5_MAV".ADDRES_22 := "P_MAV_PROFIBUS_22":P;
END_REGION

REGION Network 22: MAIN ACTUAL VALUE / FEEDBACK SPEED ADDRES 23
   RUNG wire#powerrail
      { S7_GenerateENO := "TRUE" } Move(in := "P_MAV_PROFIBUS_23":P, out1 => "DB5_MAV".ADDRES_23)
   END_RUNG
   // the same network as SCL:
   "DB5_MAV".ADDRES_23 := "P_MAV_PROFIBUS_23":P;
END_REGION

REGION Network 23: Control Word Address 2
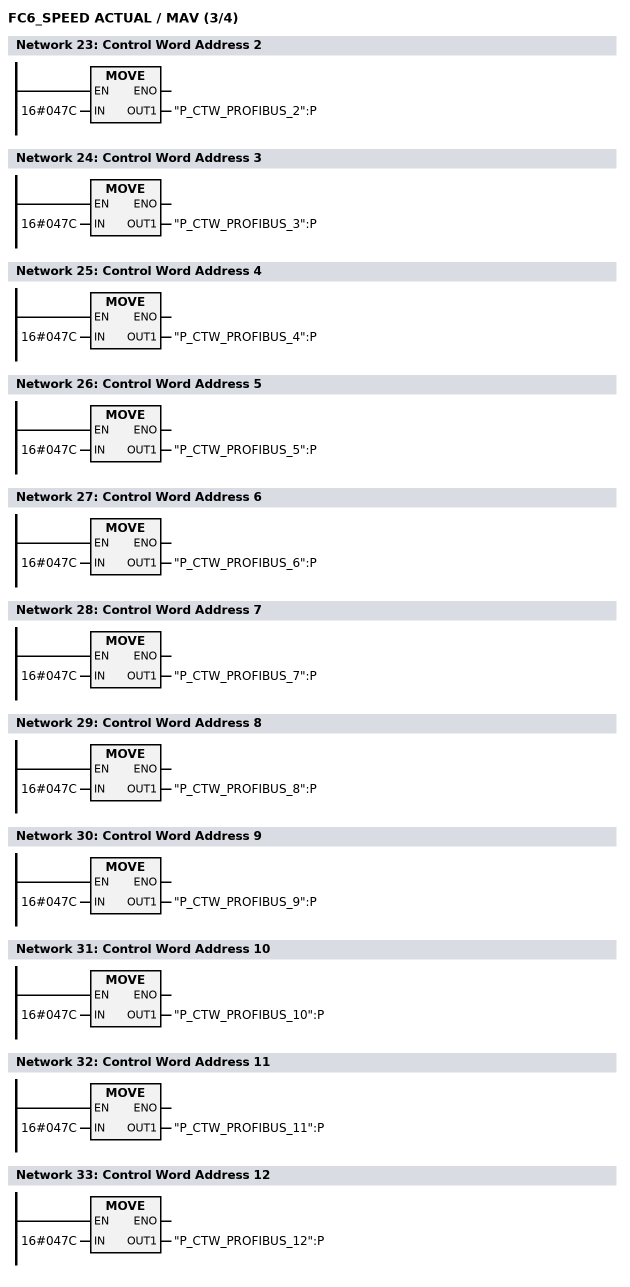
   RUNG wire#powerrail
      { S7_GenerateENO := "TRUE" } Move(in := 16#047C, out1 => "P_CTW_PROFIBUS_2":P)
   END_RUNG
   // the same network as SCL:
   "P_CTW_PROFIBUS_2":P := 16#047C;
END_REGION

REGION Network 24: Control Word Address 3
   RUNG wire#powerrail
      { S7_GenerateENO := "TRUE" } Move(in := 16#047C, out1 => "P_CTW_PROFIBUS_3":P)
   END_RUNG
   // the same network as SCL:
   "P_CTW_PROFIBUS_3":P := 16#047C;
END_REGION

REGION Network 25: Control Word Address 4
   RUNG wire#powerrail
      { S7_GenerateENO := "TRUE" } Move(in := 16#047C, out1 => "P_CTW_PROFIBUS_4":P)
   END_RUNG
   // the same network as SCL:
   "P_CTW_PROFIBUS_4":P := 16#047C;
END_REGION

REGION Network 26: Control Word Address 5
   RUNG wire#powerrail
      { S7_GenerateENO := "TRUE" } Move(in := 16#047C, out1 => "P_CTW_PROFIBUS_5":P)
   END_RUNG
   // the same network as SCL:
   "P_CTW_PROFIBUS_5":P := 16#047C;
END_REGION

REGION Network 27: Control Word Address 6
   RUNG wire#powerrail
      { S7_GenerateENO := "TRUE" } Move(in := 16#047C, out1 => "P_CTW_PROFIBUS_6":P)
   END_RUNG
   // the same network as SCL:
   "P_CTW_PROFIBUS_6":P := 16#047C;
END_REGION

REGION Network 28: Control Word Address 7
   RUNG wire#powerrail
      { S7_GenerateENO := "TRUE" } Move(in := 16#047C, out1 => "P_CTW_PROFIBUS_7":P)
   END_RUNG
   // the same network as SCL:
   "P_CTW_PROFIBUS_7":P := 16#047C;
END_REGION

REGION Network 29: Control Word Address 8
   RUNG wire#powerrail
      { S7_GenerateENO := "TRUE" } Move(in := 16#047C, out1 => "P_CTW_PROFIBUS_8":P)
   END_RUNG
   // the same network as SCL:
   "P_CTW_PROFIBUS_8":P := 16#047C;
END_REGION

REGION Network 30: Control Word Address 9
   RUNG wire#powerrail
      { S7_GenerateENO := "TRUE" } Move(in := 16#047C, out1 => "P_CTW_PROFIBUS_9":P)
   END_RUNG
   // the same network as SCL:
   "P_CTW_PROFIBUS_9":P := 16#047C;
END_REGION

REGION Network 31: Control Word Address 10
   RUNG wire#powerrail
      { S7_GenerateENO := "TRUE" } Move(in := 16#047C, out1 => "P_CTW_PROFIBUS_10":P)
   END_RUNG
   // the same network as SCL:
   "P_CTW_PROFIBUS_10":P := 16#047C;
END_REGION

REGION Network 32: Control Word Address 11
   RUNG wire#powerrail
      { S7_GenerateENO := "TRUE" } Move(in := 16#047C, out1 => "P_CTW_PROFIBUS_11":P)
   END_RUNG
   // the same network as SCL:
   "P_CTW_PROFIBUS_11":P := 16#047C;
END_REGION
